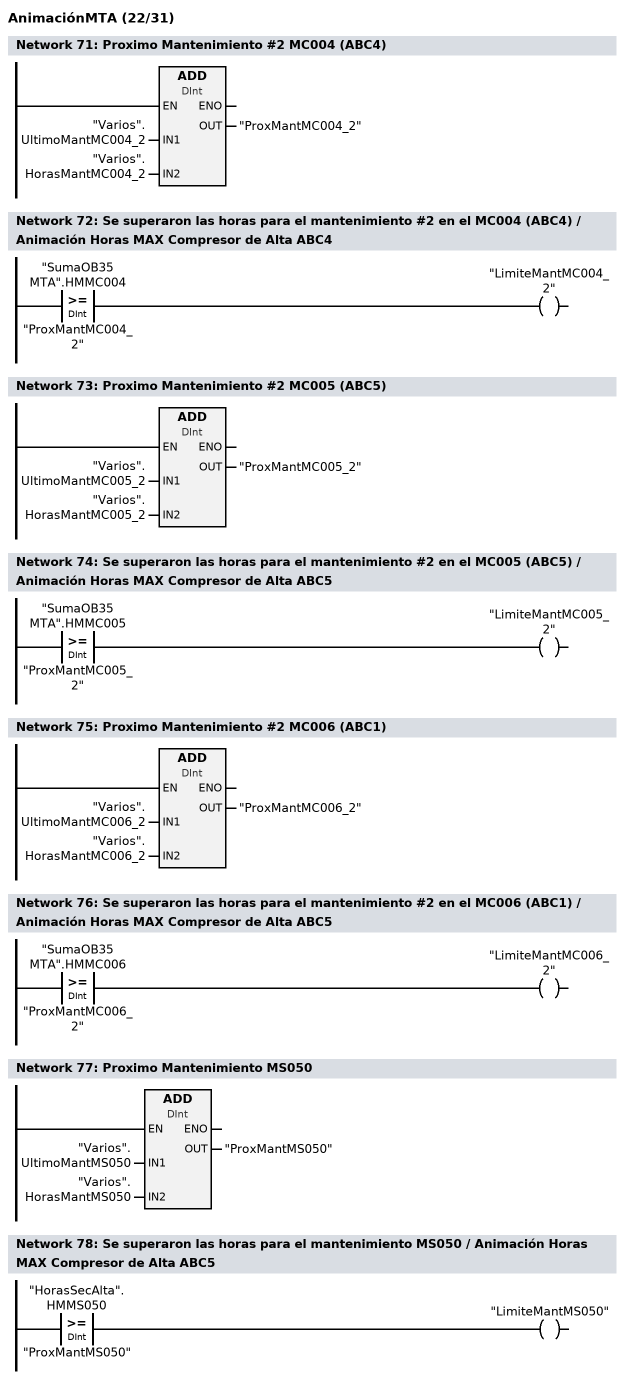
   RUNG wire#powerrail
      { S7_Templates := "SrcType := DInt"; S7_GenerateENO := "TRUE" } Add(in1 := "Varios".UltimoMantMC004_2, in2 := "Varios".HorasMantMC004_2, out => "ProxMantMC004_2")
   END_RUNG
   // the same network as SCL:
   "ProxMantMC004_2" := "Varios".UltimoMantMC004_2 + "Varios".HorasMantMC004_2;
END_REGION

REGION Network 72: Se superaron las horas para el mantenimiento #2 en el MC004 (ABC4) / Animación Horas MAX Compresor de Alta ABC4
   RUNG wire#powerrail
      { S7_Templates := "SrcType := DInt" } GE_Contact(in1 := "SumaOB35 MTA".HMMC004, in2 := "ProxMantMC004_2")
      Coil( "LimiteMantMC004_2" )
   END_RUNG
   // the same network as SCL:
   "LimiteMantMC004_2" := "SumaOB35 MTA".HMMC004 >= "ProxMantMC004_2";
END_REGION

REGION Network 73: Proximo Mantenimiento #2 MC005 (ABC5)
   RUNG wire#powerrail
      { S7_Templates := "SrcType := DInt"; S7_GenerateENO := "TRUE" } Add(in1 := "Varios".UltimoMantMC005_2, in2 := "Varios".HorasMantMC005_2, out => "ProxMantMC005_2")
   END_RUNG
   // the same network as SCL:
   "ProxMantMC005_2" := "Varios".UltimoMantMC005_2 + "Varios".HorasMantMC005_2;
END_REGION

REGION Network 74: Se superaron las horas para el mantenimiento #2 en el MC005 (ABC5) / Animación Horas MAX Compresor de Alta ABC5
   RUNG wire#powerrail
      { S7_Templates := "SrcType := DInt" } GE_Contact(in1 := "SumaOB35 MTA".HMMC005, in2 := "ProxMantMC005_2")
      Coil( "LimiteMantMC005_2" )
   END_RUNG
   // the same network as SCL:
   "LimiteMantMC005_2" := "SumaOB35 MTA".HMMC005 >= "ProxMantMC005_2";
END_REGION

REGION Network 75: Proximo Mantenimiento #2 MC006 (ABC1)
   RUNG wire#powerrail
      { S7_Templates := "SrcType := DInt"; S7_GenerateENO := "TRUE" } Add(in1 := "Varios".UltimoMantMC006_2, in2 := "Varios".HorasMantMC006_2, out => "ProxMantMC006_2")
   END_RUNG
   // the same network as SCL:
   "ProxMantMC006_2" := "Varios".UltimoMantMC006_2 + "Varios".HorasMantMC006_2;
END_REGION

REGION Network 76: Se superaron las horas para el mantenimiento #2 en el MC006 (ABC1) / Animación Horas MAX Compresor de Alta ABC5
   RUNG wire#powerrail
      { S7_Templates := "SrcType := DInt" } GE_Contact(in1 := "SumaOB35 MTA".HMMC006, in2 := "ProxMantMC006_2")
      Coil( "LimiteMantMC006_2" )
   END_RUNG
   // the same network as SCL:
   "LimiteMantMC006_2" := "SumaOB35 MTA".HMMC006 >= "ProxMantMC006_2";
END_REGION

REGION Network 77: Proximo Mantenimiento MS050
   RUNG wire#powerrail
      { S7_Templates := "SrcType := DInt"; S7_GenerateENO := "TRUE" } Add(in1 := "Varios".UltimoMantMS050, in2 := "Varios".HorasMantMS050, out => "ProxMantMS050")
   END_RUNG
   // the same network as SCL:
   "ProxMantMS050" := "Varios".UltimoMantMS050 + "Varios".HorasMantMS050;
END_REGION

REGION Network 78: Se superaron las horas para el mantenimiento MS050 / Animación Horas MAX Compresor de Alta ABC5
   RUNG wire#powerrail
      { S7_Templates := "SrcType := DInt" } GE_Contact(in1 := "HorasSecAlta".HMMS050, in2 := "ProxMantMS050")
      Coil( "LimiteMantMS050" )
   END_RUNG
   // the same network as SCL:
   "LimiteMantMS050" := "HorasSecAlta".HMMS050 >= "ProxMantMS050";
END_REGION

REGION Network 79: Proximo Mantenimiento MS051
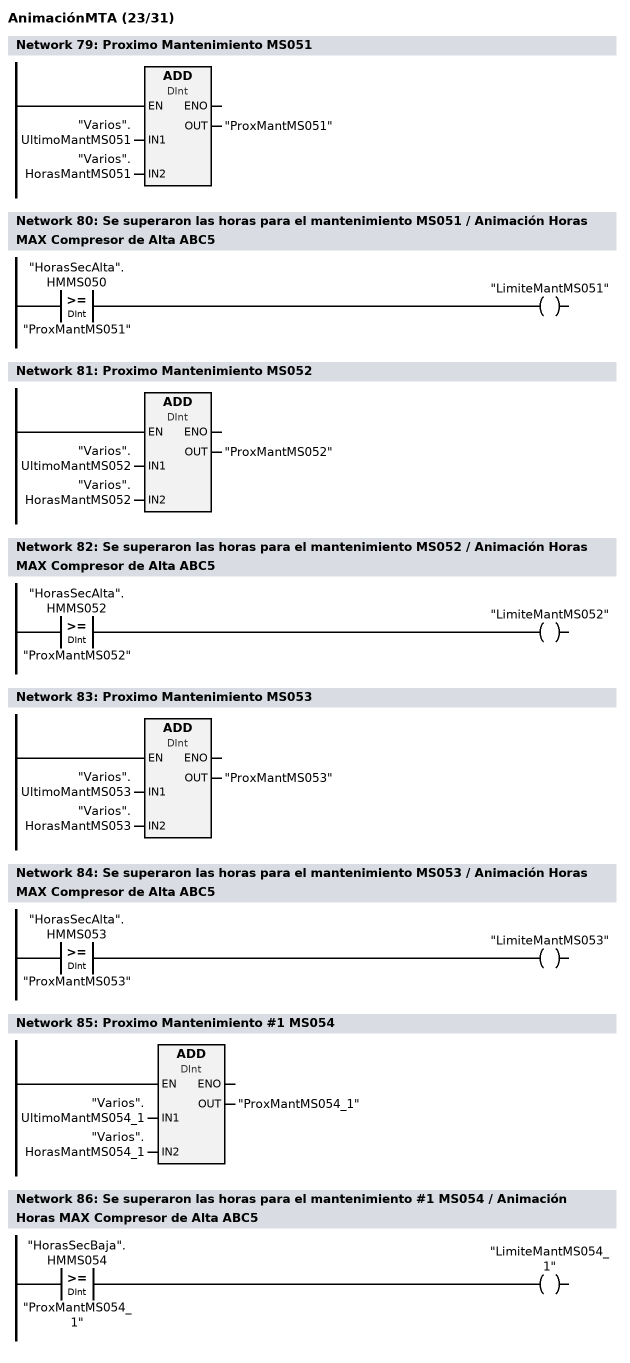
   RUNG wire#powerrail
      { S7_Templates := "SrcType := DInt"; S7_GenerateENO := "TRUE" } Add(in1 := "Varios".UltimoMantMS051, in2 := "Varios".HorasMantMS051, out => "ProxMantMS051")
   END_RUNG
   // the same network as SCL:
   "ProxMantMS051" := "Varios".UltimoMantMS051 + "Varios".HorasMantMS051;
END_REGION

REGION Network 80: Se superaron las horas para el mantenimiento MS051 / Animación Horas MAX Compresor de Alta ABC5
   RUNG wire#powerrail
      { S7_Templates := "SrcType := DInt" } GE_Contact(in1 := "HorasSecAlta".HMMS050, in2 := "ProxMantMS051")
      Coil( "LimiteMantMS051" )
   END_RUNG
   // the same network as SCL:
   "LimiteMantMS051" := "HorasSecAlta".HMMS050 >= "ProxMantMS051";
END_REGION

REGION Network 81: Proximo Mantenimiento MS052
   RUNG wire#powerrail
      { S7_Templates := "SrcType := DInt"; S7_GenerateENO := "TRUE" } Add(in1 := "Varios".UltimoMantMS052, in2 := "Varios".HorasMantMS052, out => "ProxMantMS052")
   END_RUNG
   // the same network as SCL:
   "ProxMantMS052" := "Varios".UltimoMantMS052 + "Varios".HorasMantMS052;
END_REGION

REGION Network 82: Se superaron las horas para el mantenimiento MS052 / Animación Horas MAX Compresor de Alta ABC5
   RUNG wire#powerrail
      { S7_Templates := "SrcType := DInt" } GE_Contact(in1 := "HorasSecAlta".HMMS052, in2 := "ProxMantMS052")
      Coil( "LimiteMantMS052" )
   END_RUNG
   // the same network as SCL:
   "LimiteMantMS052" := "HorasSecAlta".HMMS052 >= "ProxMantMS052";
END_REGION

REGION Network 83: Proximo Mantenimiento MS053
   RUNG wire#powerrail
      { S7_Templates := "SrcType := DInt"; S7_GenerateENO := "TRUE" } Add(in1 := "Varios".UltimoMantMS053, in2 := "Varios".HorasMantMS053, out => "ProxMantMS053")
   END_RUNG
   // the same network as SCL:
   "ProxMantMS053" := "Varios".UltimoMantMS053 + "Varios".HorasMantMS053;
END_REGION

REGION Network 84: Se superaron las horas para el mantenimiento MS053 / Animación Horas MAX Compresor de Alta ABC5
   RUNG wire#powerrail
      { S7_Templates := "SrcType := DInt" } GE_Contact(in1 := "HorasSecAlta".HMMS053, in2 := "ProxMantMS053")
      Coil( "LimiteMantMS053" )
   END_RUNG
   // the same network as SCL:
   "LimiteMantMS053" := "HorasSecAlta".HMMS053 >= "ProxMantMS053";
END_REGION

REGION Network 85: Proximo Mantenimiento #1 MS054
   RUNG wire#powerrail
      { S7_Templates := "SrcType := DInt"; S7_GenerateENO := "TRUE" } Add(in1 := "Varios".UltimoMantMS054_1, in2 := "Varios".HorasMantMS054_1, out => "ProxMantMS054_1")
   END_RUNG
   // the same network as SCL:
   "ProxMantMS054_1" := "Varios".UltimoMantMS054_1 + "Varios".HorasMantMS054_1;
END_REGION

REGION Network 86: Se superaron las horas para el mantenimiento #1 MS054 / Animación Horas MAX Compresor de Alta ABC5
   RUNG wire#powerrail
      { S7_Templates := "SrcType := DInt" } GE_Contact(in1 := "HorasSecBaja".HMMS054, in2 := "ProxMantMS054_1")
      Coil( "LimiteMantMS054_1" )
   END_RUNG
   // the same network as SCL:
   "LimiteMantMS054_1" := "HorasSecBaja".HMMS054 >= "ProxMantMS054_1";
END_REGION

REGION Network 87: Proximo Mantenimiento #2 MS054
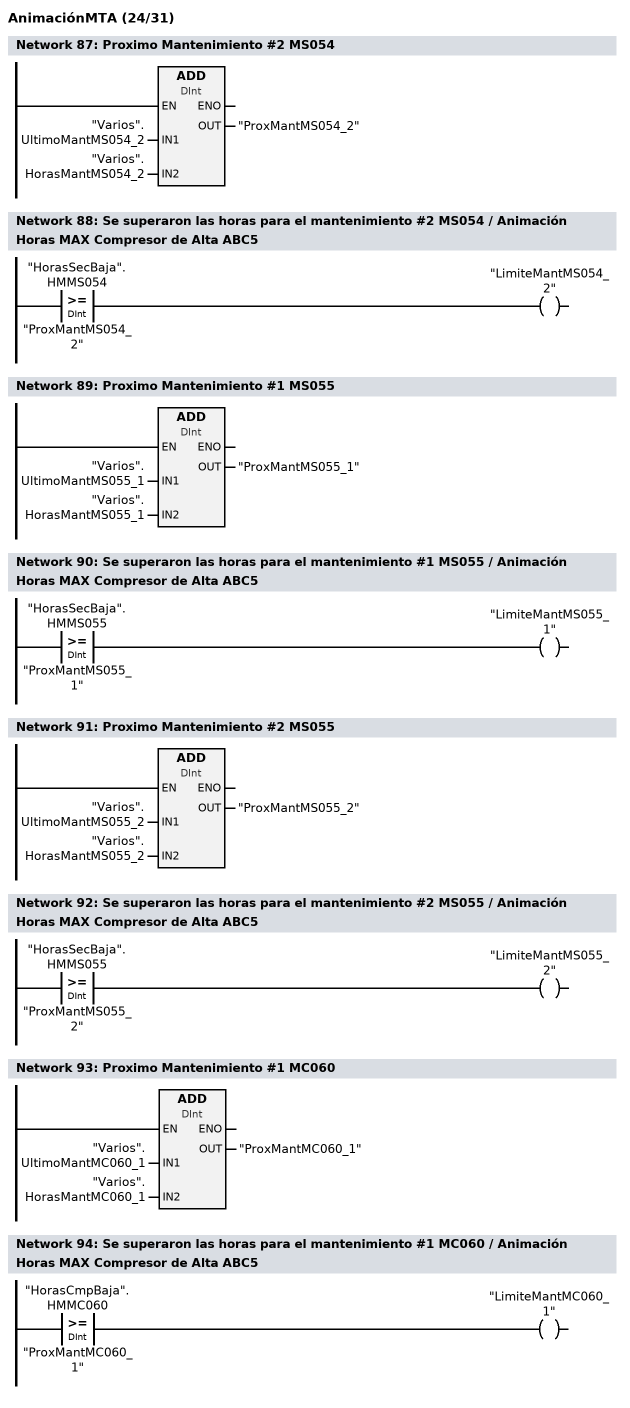
   RUNG wire#powerrail
      { S7_Templates := "SrcType := DInt"; S7_GenerateENO := "TRUE" } Add(in1 := "Varios".UltimoMantMS054_2, in2 := "Varios".HorasMantMS054_2, out => "ProxMantMS054_2")
   END_RUNG
   // the same network as SCL:
   "ProxMantMS054_2" := "Varios".UltimoMantMS054_2 + "Varios".HorasMantMS054_2;
END_REGION

REGION Network 88: Se superaron las horas para el mantenimiento #2 MS054 / Animación Horas MAX Compresor de Alta ABC5
   RUNG wire#powerrail
      { S7_Templates := "SrcType := DInt" } GE_Contact(in1 := "HorasSecBaja".HMMS054, in2 := "ProxMantMS054_2")
      Coil( "LimiteMantMS054_2" )
   END_RUNG
   // the same network as SCL:
   "LimiteMantMS054_2" := "HorasSecBaja".HMMS054 >= "ProxMantMS054_2";
END_REGION

REGION Network 89: Proximo Mantenimiento #1 MS055
   RUNG wire#powerrail
      { S7_Templates := "SrcType := DInt"; S7_GenerateENO := "TRUE" } Add(in1 := "Varios".UltimoMantMS055_1, in2 := "Varios".HorasMantMS055_1, out => "ProxMantMS055_1")
   END_RUNG
   // the same network as SCL:
   "ProxMantMS055_1" := "Varios".UltimoMantMS055_1 + "Varios".HorasMantMS055_1;
END_REGION

REGION Network 90: Se superaron las horas para el mantenimiento #1 MS055 / Animación Horas MAX Compresor de Alta ABC5
   RUNG wire#powerrail
      { S7_Templates := "SrcType := DInt" } GE_Contact(in1 := "HorasSecBaja".HMMS055, in2 := "ProxMantMS055_1")
      Coil( "LimiteMantMS055_1" )
   END_RUNG
   // the same network as SCL:
   "LimiteMantMS055_1" := "HorasSecBaja".HMMS055 >= "ProxMantMS055_1";
END_REGION

REGION Network 91: Proximo Mantenimiento #2 MS055
   RUNG wire#powerrail
      { S7_Templates := "SrcType := DInt"; S7_GenerateENO := "TRUE" } Add(in1 := "Varios".UltimoMantMS055_2, in2 := "Varios".HorasMantMS055_2, out => "ProxMantMS055_2")
   END_RUNG
   // the same network as SCL:
   "ProxMantMS055_2" := "Varios".UltimoMantMS055_2 + "Varios".HorasMantMS055_2;
END_REGION

REGION Network 92: Se superaron las horas para el mantenimiento #2 MS055 / Animación Horas MAX Compresor de Alta ABC5
   RUNG wire#powerrail
      { S7_Templates := "SrcType := DInt" } GE_Contact(in1 := "HorasSecBaja".HMMS055, in2 := "ProxMantMS055_2")
      Coil( "LimiteMantMS055_2" )
   END_RUNG
   // the same network as SCL:
   "LimiteMantMS055_2" := "HorasSecBaja".HMMS055 >= "ProxMantMS055_2";
END_REGION

REGION Network 93: Proximo Mantenimiento #1 MC060
   RUNG wire#powerrail
      { S7_Templates := "SrcType := DInt"; S7_GenerateENO := "TRUE" } Add(in1 := "Varios".UltimoMantMC060_1, in2 := "Varios".HorasMantMC060_1, out => "ProxMantMC060_1")
   END_RUNG
   // the same network as SCL:
   "ProxMantMC060_1" := "Varios".UltimoMantMC060_1 + "Varios".HorasMantMC060_1;
END_REGION

REGION Network 94: Se superaron las horas para el mantenimiento #1 MC060 / Animación Horas MAX Compresor de Alta ABC5
   RUNG wire#powerrail
      { S7_Templates := "SrcType := DInt" } GE_Contact(in1 := "HorasCmpBaja".HMMC060, in2 := "ProxMantMC060_1")
      Coil( "LimiteMantMC060_1" )
   END_RUNG
   // the same network as SCL:
   "LimiteMantMC060_1" := "HorasCmpBaja".HMMC060 >= "ProxMantMC060_1";
END_REGION

REGION Network 95: Proximo Mantenimiento #2 MC060
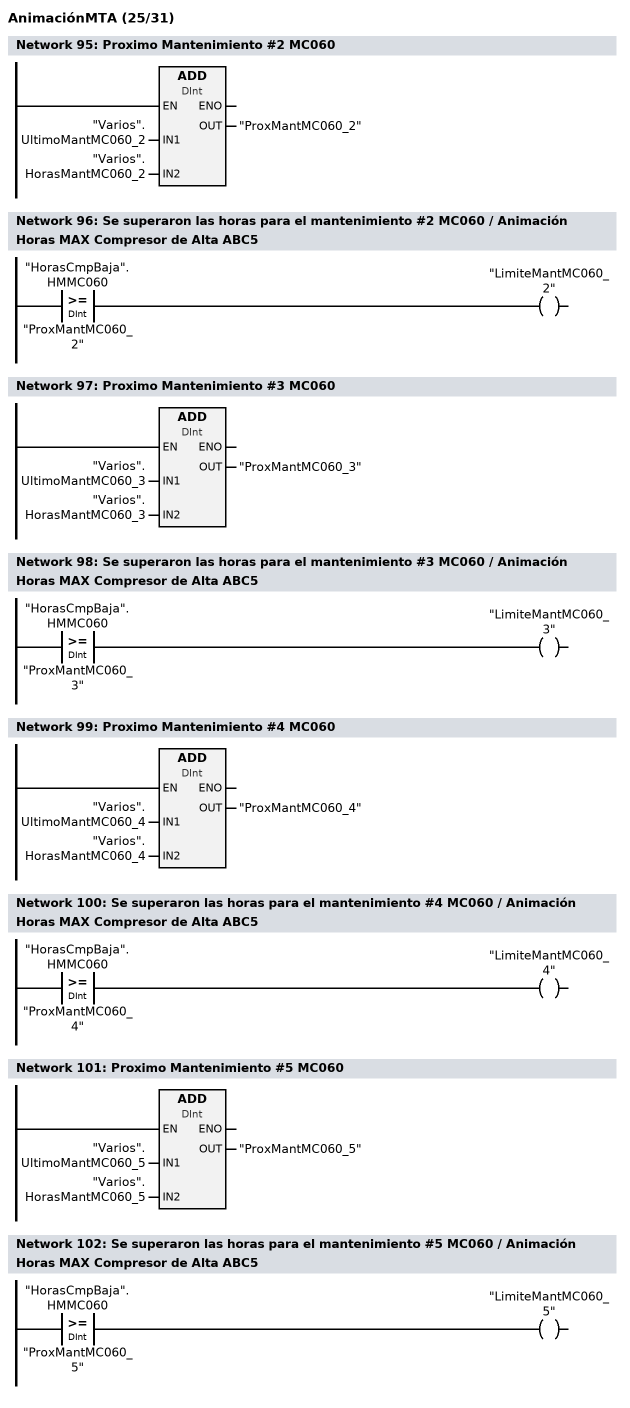
   RUNG wire#powerrail
      { S7_Templates := "SrcType := DInt"; S7_GenerateENO := "TRUE" } Add(in1 := "Varios".UltimoMantMC060_2, in2 := "Varios".HorasMantMC060_2, out => "ProxMantMC060_2")
   END_RUNG
   // the same network as SCL:
   "ProxMantMC060_2" := "Varios".UltimoMantMC060_2 + "Varios".HorasMantMC060_2;
END_REGION

REGION Network 96: Se superaron las horas para el mantenimiento #2 MC060 / Animación Horas MAX Compresor de Alta ABC5
   RUNG wire#powerrail
      { S7_Templates := "SrcType := DInt" } GE_Contact(in1 := "HorasCmpBaja".HMMC060, in2 := "ProxMantMC060_2")
      Coil( "LimiteMantMC060_2" )
   END_RUNG
   // the same network as SCL:
   "LimiteMantMC060_2" := "HorasCmpBaja".HMMC060 >= "ProxMantMC060_2";
END_REGION

REGION Network 97: Proximo Mantenimiento #3 MC060
   RUNG wire#powerrail
      { S7_Templates := "SrcType := DInt"; S7_GenerateENO := "TRUE" } Add(in1 := "Varios".UltimoMantMC060_3, in2 := "Varios".HorasMantMC060_3, out => "ProxMantMC060_3")
   END_RUNG
   // the same network as SCL:
   "ProxMantMC060_3" := "Varios".UltimoMantMC060_3 + "Varios".HorasMantMC060_3;
END_REGION

REGION Network 98: Se superaron las horas para el mantenimiento #3 MC060 / Animación Horas MAX Compresor de Alta ABC5
   RUNG wire#powerrail
      { S7_Templates := "SrcType := DInt" } GE_Contact(in1 := "HorasCmpBaja".HMMC060, in2 := "ProxMantMC060_3")
      Coil( "LimiteMantMC060_3" )
   END_RUNG
   // the same network as SCL:
   "LimiteMantMC060_3" := "HorasCmpBaja".HMMC060 >= "ProxMantMC060_3";
END_REGION

REGION Network 99: Proximo Mantenimiento #4 MC060
   RUNG wire#powerrail
      { S7_Templates := "SrcType := DInt"; S7_GenerateENO := "TRUE" } Add(in1 := "Varios".UltimoMantMC060_4, in2 := "Varios".HorasMantMC060_4, out => "ProxMantMC060_4")
   END_RUNG
   // the same network as SCL:
   "ProxMantMC060_4" := "Varios".UltimoMantMC060_4 + "Varios".HorasMantMC060_4;
END_REGION

REGION Network 100: Se superaron las horas para el mantenimiento #4 MC060 / Animación Horas MAX Compresor de Alta ABC5
   RUNG wire#powerrail
      { S7_Templates := "SrcType := DInt" } GE_Contact(in1 := "HorasCmpBaja".HMMC060, in2 := "ProxMantMC060_4")
      Coil( "LimiteMantMC060_4" )
   END_RUNG
   // the same network as SCL:
   "LimiteMantMC060_4" := "HorasCmpBaja".HMMC060 >= "ProxMantMC060_4";
END_REGION

REGION Network 101: Proximo Mantenimiento #5 MC060
   RUNG wire#powerrail
      { S7_Templates := "SrcType := DInt"; S7_GenerateENO := "TRUE" } Add(in1 := "Varios".UltimoMantMC060_5, in2 := "Varios".HorasMantMC060_5, out => "ProxMantMC060_5")
   END_RUNG
   // the same network as SCL:
   "ProxMantMC060_5" := "Varios".UltimoMantMC060_5 + "Varios".HorasMantMC060_5;
END_REGION

REGION Network 102: Se superaron las horas para el mantenimiento #5 MC060 / Animación Horas MAX Compresor de Alta ABC5
   RUNG wire#powerrail
      { S7_Templates := "SrcType := DInt" } GE_Contact(in1 := "HorasCmpBaja".HMMC060, in2 := "ProxMantMC060_5")
      Coil( "LimiteMantMC060_5" )
   END_RUNG
   // the same network as SCL:
   "LimiteMantMC060_5" := "HorasCmpBaja".HMMC060 >= "ProxMantMC060_5";
END_REGION

REGION Network 103: Proximo Mantenimiento #1 MC061
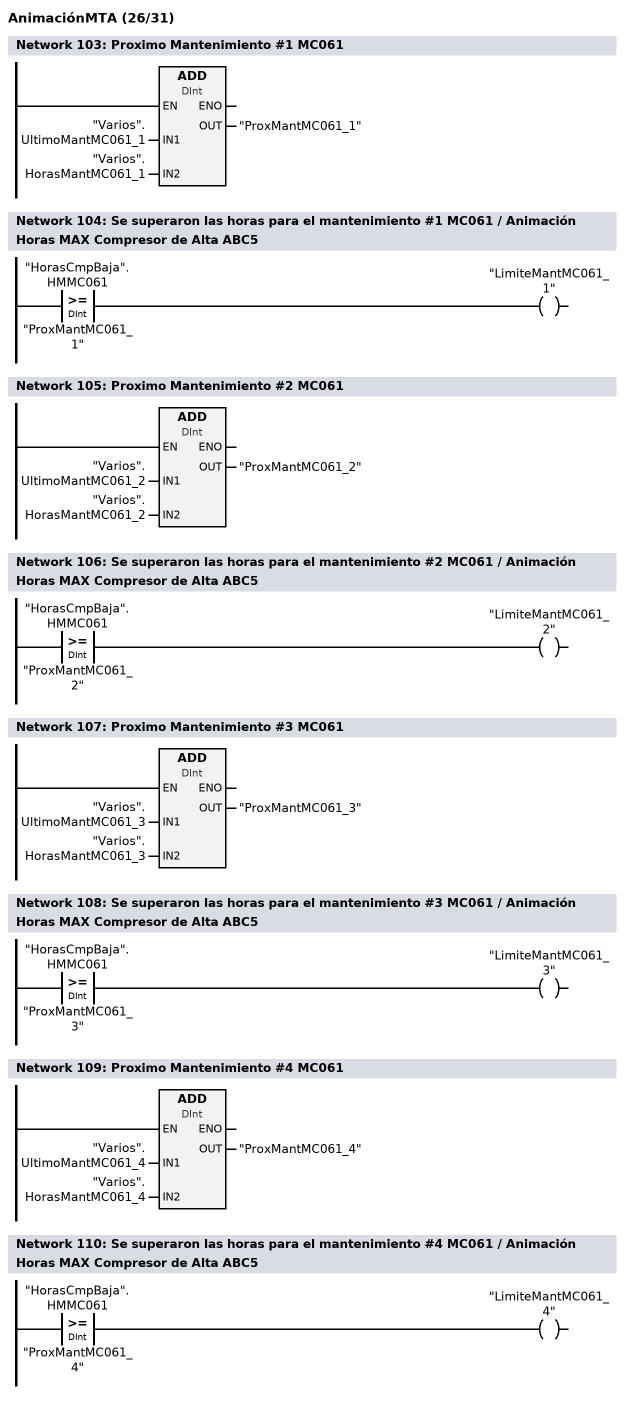
   RUNG wire#powerrail
      { S7_Templates := "SrcType := DInt"; S7_GenerateENO := "TRUE" } Add(in1 := "Varios".UltimoMantMC061_1, in2 := "Varios".HorasMantMC061_1, out => "ProxMantMC061_1")
   END_RUNG
   // the same network as SCL:
   "ProxMantMC061_1" := "Varios".UltimoMantMC061_1 + "Varios".HorasMantMC061_1;
END_REGION

REGION Network 104: Se superaron las horas para el mantenimiento #1 MC061 / Animación Horas MAX Compresor de Alta ABC5
   RUNG wire#powerrail
      { S7_Templates := "SrcType := DInt" } GE_Contact(in1 := "HorasCmpBaja".HMMC061, in2 := "ProxMantMC061_1")
      Coil( "LimiteMantMC061_1" )
   END_RUNG
   // the same network as SCL:
   "LimiteMantMC061_1" := "HorasCmpBaja".HMMC061 >= "ProxMantMC061_1";
END_REGION

REGION Network 105: Proximo Mantenimiento #2 MC061
   RUNG wire#powerrail
      { S7_Templates := "SrcType := DInt"; S7_GenerateENO := "TRUE" } Add(in1 := "Varios".UltimoMantMC061_2, in2 := "Varios".HorasMantMC061_2, out => "ProxMantMC061_2")
   END_RUNG
   // the same network as SCL:
   "ProxMantMC061_2" := "Varios".UltimoMantMC061_2 + "Varios".HorasMantMC061_2;
END_REGION

REGION Network 106: Se superaron las horas para el mantenimiento #2 MC061 / Animación Horas MAX Compresor de Alta ABC5
   RUNG wire#powerrail
      { S7_Templates := "SrcType := DInt" } GE_Contact(in1 := "HorasCmpBaja".HMMC061, in2 := "ProxMantMC061_2")
      Coil( "LimiteMantMC061_2" )
   END_RUNG
   // the same network as SCL:
   "LimiteMantMC061_2" := "HorasCmpBaja".HMMC061 >= "ProxMantMC061_2";
END_REGION

REGION Network 107: Proximo Mantenimiento #3 MC061
   RUNG wire#powerrail
      { S7_Templates := "SrcType := DInt"; S7_GenerateENO := "TRUE" } Add(in1 := "Varios".UltimoMantMC061_3, in2 := "Varios".HorasMantMC061_3, out => "ProxMantMC061_3")
   END_RUNG
   // the same network as SCL:
   "ProxMantMC061_3" := "Varios".UltimoMantMC061_3 + "Varios".HorasMantMC061_3;
END_REGION

REGION Network 108: Se superaron las horas para el mantenimiento #3 MC061 / Animación Horas MAX Compresor de Alta ABC5
   RUNG wire#powerrail
      { S7_Templates := "SrcType := DInt" } GE_Contact(in1 := "HorasCmpBaja".HMMC061, in2 := "ProxMantMC061_3")
      Coil( "LimiteMantMC061_3" )
   END_RUNG
   // the same network as SCL:
   "LimiteMantMC061_3" := "HorasCmpBaja".HMMC061 >= "ProxMantMC061_3";
END_REGION

REGION Network 109: Proximo Mantenimiento #4 MC061
   RUNG wire#powerrail
      { S7_Templates := "SrcType := DInt"; S7_GenerateENO := "TRUE" } Add(in1 := "Varios".UltimoMantMC061_4, in2 := "Varios".HorasMantMC061_4, out => "ProxMantMC061_4")
   END_RUNG
   // the same network as SCL:
   "ProxMantMC061_4" := "Varios".UltimoMantMC061_4 + "Varios".HorasMantMC061_4;
END_REGION

REGION Network 110: Se superaron las horas para el mantenimiento #4 MC061 / Animación Horas MAX Compresor de Alta ABC5
   RUNG wire#powerrail
      { S7_Templates := "SrcType := DInt" } GE_Contact(in1 := "HorasCmpBaja".HMMC061, in2 := "ProxMantMC061_4")
      Coil( "LimiteMantMC061_4" )
   END_RUNG
   // the same network as SCL:
   "LimiteMantMC061_4" := "HorasCmpBaja".HMMC061 >= "ProxMantMC061_4";
END_REGION

REGION Network 111: Proximo Mantenimiento #5 MC061
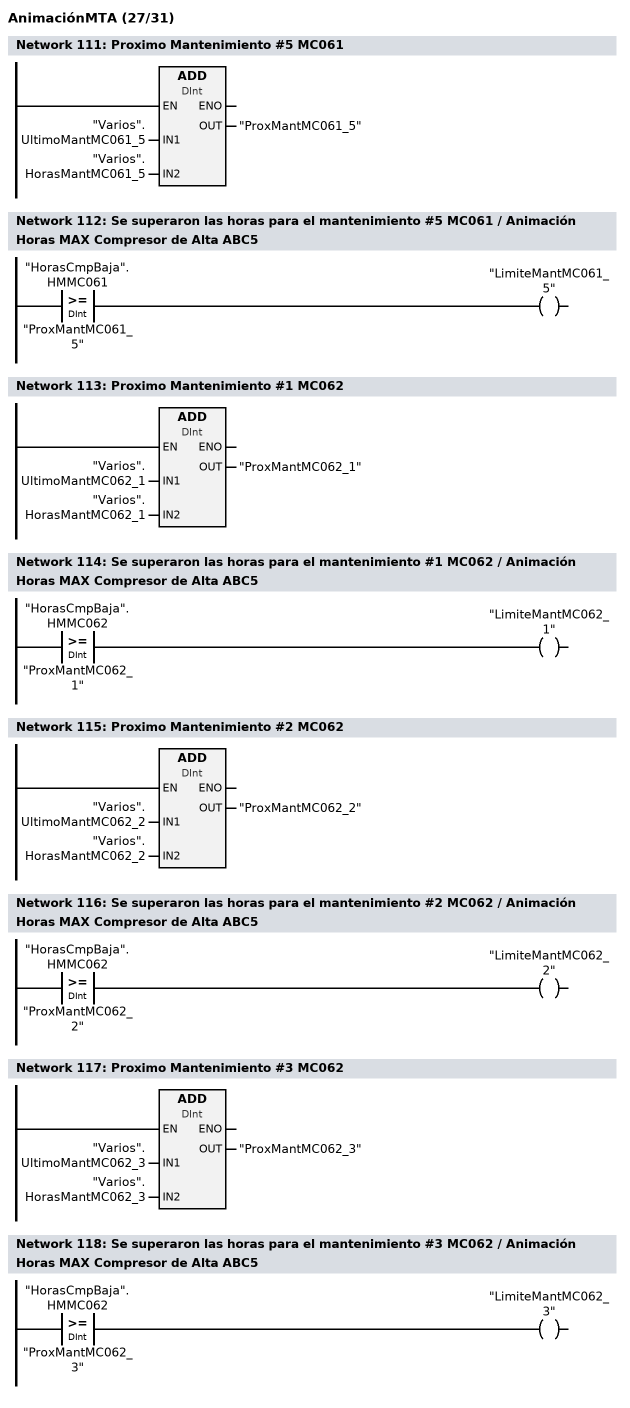
   RUNG wire#powerrail
      { S7_Templates := "SrcType := DInt"; S7_GenerateENO := "TRUE" } Add(in1 := "Varios".UltimoMantMC061_5, in2 := "Varios".HorasMantMC061_5, out => "ProxMantMC061_5")
   END_RUNG
   // the same network as SCL:
   "ProxMantMC061_5" := "Varios".UltimoMantMC061_5 + "Varios".HorasMantMC061_5;
END_REGION

REGION Network 112: Se superaron las horas para el mantenimiento #5 MC061 / Animación Horas MAX Compresor de Alta ABC5
   RUNG wire#powerrail
      { S7_Templates := "SrcType := DInt" } GE_Contact(in1 := "HorasCmpBaja".HMMC061, in2 := "ProxMantMC061_5")
      Coil( "LimiteMantMC061_5" )
   END_RUNG
   // the same network as SCL:
   "LimiteMantMC061_5" := "HorasCmpBaja".HMMC061 >= "ProxMantMC061_5";
END_REGION

REGION Network 113: Proximo Mantenimiento #1 MC062
   RUNG wire#powerrail
      { S7_Templates := "SrcType := DInt"; S7_GenerateENO := "TRUE" } Add(in1 := "Varios".UltimoMantMC062_1, in2 := "Varios".HorasMantMC062_1, out => "ProxMantMC062_1")
   END_RUNG
   // the same network as SCL:
   "ProxMantMC062_1" := "Varios".UltimoMantMC062_1 + "Varios".HorasMantMC062_1;
END_REGION

REGION Network 114: Se superaron las horas para el mantenimiento #1 MC062 / Animación Horas MAX Compresor de Alta ABC5
   RUNG wire#powerrail
      { S7_Templates := "SrcType := DInt" } GE_Contact(in1 := "HorasCmpBaja".HMMC062, in2 := "ProxMantMC062_1")
      Coil( "LimiteMantMC062_1" )
   END_RUNG
   // the same network as SCL:
   "LimiteMantMC062_1" := "HorasCmpBaja".HMMC062 >= "ProxMantMC062_1";
END_REGION

REGION Network 115: Proximo Mantenimiento #2 MC062
   RUNG wire#powerrail
      { S7_Templates := "SrcType := DInt"; S7_GenerateENO := "TRUE" } Add(in1 := "Varios".UltimoMantMC062_2, in2 := "Varios".HorasMantMC062_2, out => "ProxMantMC062_2")
   END_RUNG
   // the same network as SCL:
   "ProxMantMC062_2" := "Varios".UltimoMantMC062_2 + "Varios".HorasMantMC062_2;
END_REGION

REGION Network 116: Se superaron las horas para el mantenimiento #2 MC062 / Animación Horas MAX Compresor de Alta ABC5
   RUNG wire#powerrail
      { S7_Templates := "SrcType := DInt" } GE_Contact(in1 := "HorasCmpBaja".HMMC062, in2 := "ProxMantMC062_2")
      Coil( "LimiteMantMC062_2" )
   END_RUNG
   // the same network as SCL:
   "LimiteMantMC062_2" := "HorasCmpBaja".HMMC062 >= "ProxMantMC062_2";
END_REGION

REGION Network 117: Proximo Mantenimiento #3 MC062
   RUNG wire#powerrail
      { S7_Templates := "SrcType := DInt"; S7_GenerateENO := "TRUE" } Add(in1 := "Varios".UltimoMantMC062_3, in2 := "Varios".HorasMantMC062_3, out => "ProxMantMC062_3")
   END_RUNG
   // the same network as SCL:
   "ProxMantMC062_3" := "Varios".UltimoMantMC062_3 + "Varios".HorasMantMC062_3;
END_REGION

REGION Network 118: Se superaron las horas para el mantenimiento #3 MC062 / Animación Horas MAX Compresor de Alta ABC5
   RUNG wire#powerrail
      { S7_Templates := "SrcType := DInt" } GE_Contact(in1 := "HorasCmpBaja".HMMC062, in2 := "ProxMantMC062_3")
      Coil( "LimiteMantMC062_3" )
   END_RUNG
   // the same network as SCL:
   "LimiteMantMC062_3" := "HorasCmpBaja".HMMC062 >= "ProxMantMC062_3";
END_REGION

REGION Network 119: Proximo Mantenimiento #4 MC062
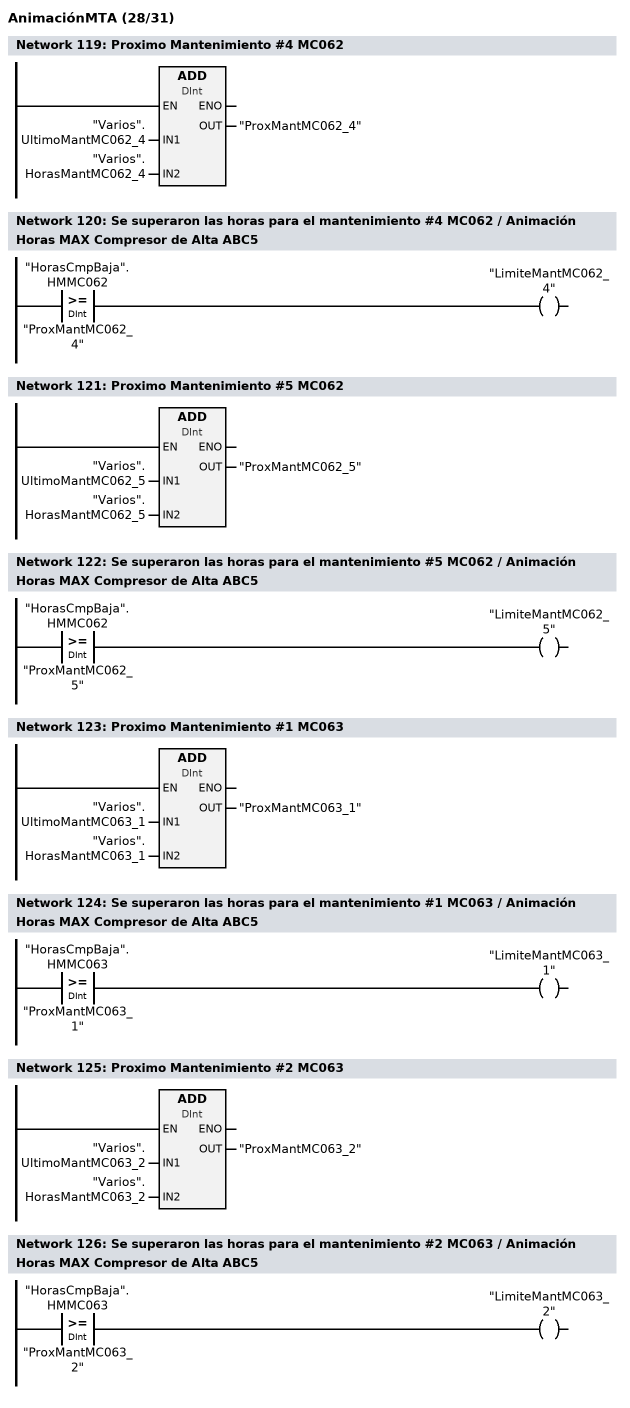
   RUNG wire#powerrail
      { S7_Templates := "SrcType := DInt"; S7_GenerateENO := "TRUE" } Add(in1 := "Varios".UltimoMantMC062_4, in2 := "Varios".HorasMantMC062_4, out => "ProxMantMC062_4")
   END_RUNG
   // the same network as SCL:
   "ProxMantMC062_4" := "Varios".UltimoMantMC062_4 + "Varios".HorasMantMC062_4;
END_REGION

REGION Network 120: Se superaron las horas para el mantenimiento #4 MC062 / Animación Horas MAX Compresor de Alta ABC5
   RUNG wire#powerrail
      { S7_Templates := "SrcType := DInt" } GE_Contact(in1 := "HorasCmpBaja".HMMC062, in2 := "ProxMantMC062_4")
      Coil( "LimiteMantMC062_4" )
   END_RUNG
   // the same network as SCL:
   "LimiteMantMC062_4" := "HorasCmpBaja".HMMC062 >= "ProxMantMC062_4";
END_REGION

REGION Network 121: Proximo Mantenimiento #5 MC062
   RUNG wire#powerrail
      { S7_Templates := "SrcType := DInt"; S7_GenerateENO := "TRUE" } Add(in1 := "Varios".UltimoMantMC062_5, in2 := "Varios".HorasMantMC062_5, out => "ProxMantMC062_5")
   END_RUNG
   // the same network as SCL:
   "ProxMantMC062_5" := "Varios".UltimoMantMC062_5 + "Varios".HorasMantMC062_5;
END_REGION

REGION Network 122: Se superaron las horas para el mantenimiento #5 MC062 / Animación Horas MAX Compresor de Alta ABC5
   RUNG wire#powerrail
      { S7_Templates := "SrcType := DInt" } GE_Contact(in1 := "HorasCmpBaja".HMMC062, in2 := "ProxMantMC062_5")
      Coil( "LimiteMantMC062_5" )
   END_RUNG
   // the same network as SCL:
   "LimiteMantMC062_5" := "HorasCmpBaja".HMMC062 >= "ProxMantMC062_5";
END_REGION

REGION Network 123: Proximo Mantenimiento #1 MC063
   RUNG wire#powerrail
      { S7_Templates := "SrcType := DInt"; S7_GenerateENO := "TRUE" } Add(in1 := "Varios".UltimoMantMC063_1, in2 := "Varios".HorasMantMC063_1, out => "ProxMantMC063_1")
   END_RUNG
   // the same network as SCL:
   "ProxMantMC063_1" := "Varios".UltimoMantMC063_1 + "Varios".HorasMantMC063_1;
END_REGION

REGION Network 124: Se superaron las horas para el mantenimiento #1 MC063 / Animación Horas MAX Compresor de Alta ABC5
   RUNG wire#powerrail
      { S7_Templates := "SrcType := DInt" } GE_Contact(in1 := "HorasCmpBaja".HMMC063, in2 := "ProxMantMC063_1")
      Coil( "LimiteMantMC063_1" )
   END_RUNG
   // the same network as SCL:
   "LimiteMantMC063_1" := "HorasCmpBaja".HMMC063 >= "ProxMantMC063_1";
END_REGION

REGION Network 125: Proximo Mantenimiento #2 MC063
   RUNG wire#powerrail
      { S7_Templates := "SrcType := DInt"; S7_GenerateENO := "TRUE" } Add(in1 := "Varios".UltimoMantMC063_2, in2 := "Varios".HorasMantMC063_2, out => "ProxMantMC063_2")
   END_RUNG
   // the same network as SCL:
   "ProxMantMC063_2" := "Varios".UltimoMantMC063_2 + "Varios".HorasMantMC063_2;
END_REGION

REGION Network 126: Se superaron las horas para el mantenimiento #2 MC063 / Animación Horas MAX Compresor de Alta ABC5
   RUNG wire#powerrail
      { S7_Templates := "SrcType := DInt" } GE_Contact(in1 := "HorasCmpBaja".HMMC063, in2 := "ProxMantMC063_2")
      Coil( "LimiteMantMC063_2" )
   END_RUNG
   // the same network as SCL:
   "LimiteMantMC063_2" := "HorasCmpBaja".HMMC063 >= "ProxMantMC063_2";
END_REGION

REGION Network 127: Proximo Mantenimiento #3 MC063
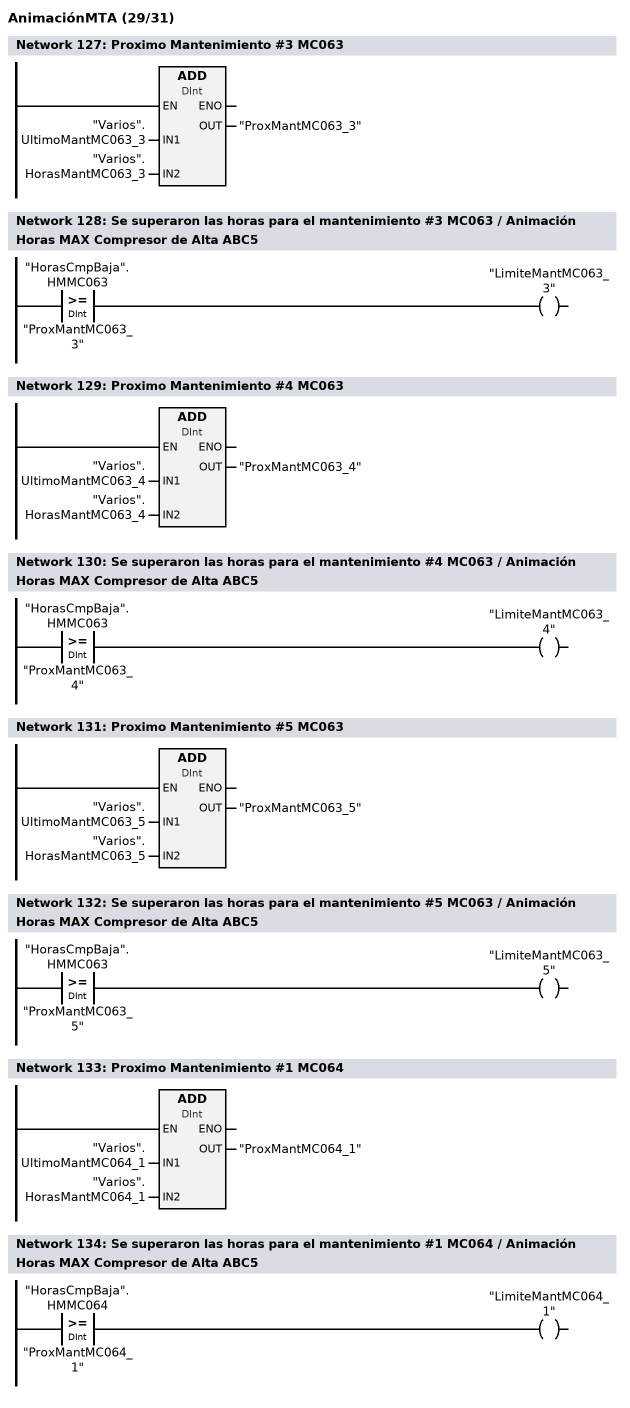
   RUNG wire#powerrail
      { S7_Templates := "SrcType := DInt"; S7_GenerateENO := "TRUE" } Add(in1 := "Varios".UltimoMantMC063_3, in2 := "Varios".HorasMantMC063_3, out => "ProxMantMC063_3")
   END_RUNG
   // the same network as SCL:
   "ProxMantMC063_3" := "Varios".UltimoMantMC063_3 + "Varios".HorasMantMC063_3;
END_REGION

REGION Network 128: Se superaron las horas para el mantenimiento #3 MC063 / Animación Horas MAX Compresor de Alta ABC5
   RUNG wire#powerrail
      { S7_Templates := "SrcType := DInt" } GE_Contact(in1 := "HorasCmpBaja".HMMC063, in2 := "ProxMantMC063_3")
      Coil( "LimiteMantMC063_3" )
   END_RUNG
   // the same network as SCL:
   "LimiteMantMC063_3" := "HorasCmpBaja".HMMC063 >= "ProxMantMC063_3";
END_REGION

REGION Network 129: Proximo Mantenimiento #4 MC063
   RUNG wire#powerrail
      { S7_Templates := "SrcType := DInt"; S7_GenerateENO := "TRUE" } Add(in1 := "Varios".UltimoMantMC063_4, in2 := "Varios".HorasMantMC063_4, out => "ProxMantMC063_4")
   END_RUNG
   // the same network as SCL:
   "ProxMantMC063_4" := "Varios".UltimoMantMC063_4 + "Varios".HorasMantMC063_4;
END_REGION

REGION Network 130: Se superaron las horas para el mantenimiento #4 MC063 / Animación Horas MAX Compresor de Alta ABC5
   RUNG wire#powerrail
      { S7_Templates := "SrcType := DInt" } GE_Contact(in1 := "HorasCmpBaja".HMMC063, in2 := "ProxMantMC063_4")
      Coil( "LimiteMantMC063_4" )
   END_RUNG
   // the same network as SCL:
   "LimiteMantMC063_4" := "HorasCmpBaja".HMMC063 >= "ProxMantMC063_4";
END_REGION

REGION Network 131: Proximo Mantenimiento #5 MC063
   RUNG wire#powerrail
      { S7_Templates := "SrcType := DInt"; S7_GenerateENO := "TRUE" } Add(in1 := "Varios".UltimoMantMC063_5, in2 := "Varios".HorasMantMC063_5, out => "ProxMantMC063_5")
   END_RUNG
   // the same network as SCL:
   "ProxMantMC063_5" := "Varios".UltimoMantMC063_5 + "Varios".HorasMantMC063_5;
END_REGION

REGION Network 132: Se superaron las horas para el mantenimiento #5 MC063 / Animación Horas MAX Compresor de Alta ABC5
   RUNG wire#powerrail
      { S7_Templates := "SrcType := DInt" } GE_Contact(in1 := "HorasCmpBaja".HMMC063, in2 := "ProxMantMC063_5")
      Coil( "LimiteMantMC063_5" )
   END_RUNG
   // the same network as SCL:
   "LimiteMantMC063_5" := "HorasCmpBaja".HMMC063 >= "ProxMantMC063_5";
END_REGION

REGION Network 133: Proximo Mantenimiento #1 MC064
   RUNG wire#powerrail
      { S7_Templates := "SrcType := DInt"; S7_GenerateENO := "TRUE" } Add(in1 := "Varios".UltimoMantMC064_1, in2 := "Varios".HorasMantMC064_1, out => "ProxMantMC064_1")
   END_RUNG
   // the same network as SCL:
   "ProxMantMC064_1" := "Varios".UltimoMantMC064_1 + "Varios".HorasMantMC064_1;
END_REGION

REGION Network 134: Se superaron las horas para el mantenimiento #1 MC064 / Animación Horas MAX Compresor de Alta ABC5
   RUNG wire#powerrail
      { S7_Templates := "SrcType := DInt" } GE_Contact(in1 := "HorasCmpBaja".HMMC064, in2 := "ProxMantMC064_1")
      Coil( "LimiteMantMC064_1" )
   END_RUNG
   // the same network as SCL:
   "LimiteMantMC064_1" := "HorasCmpBaja".HMMC064 >= "ProxMantMC064_1";
END_REGION

REGION Network 135: Proximo Mantenimiento #2 MC064
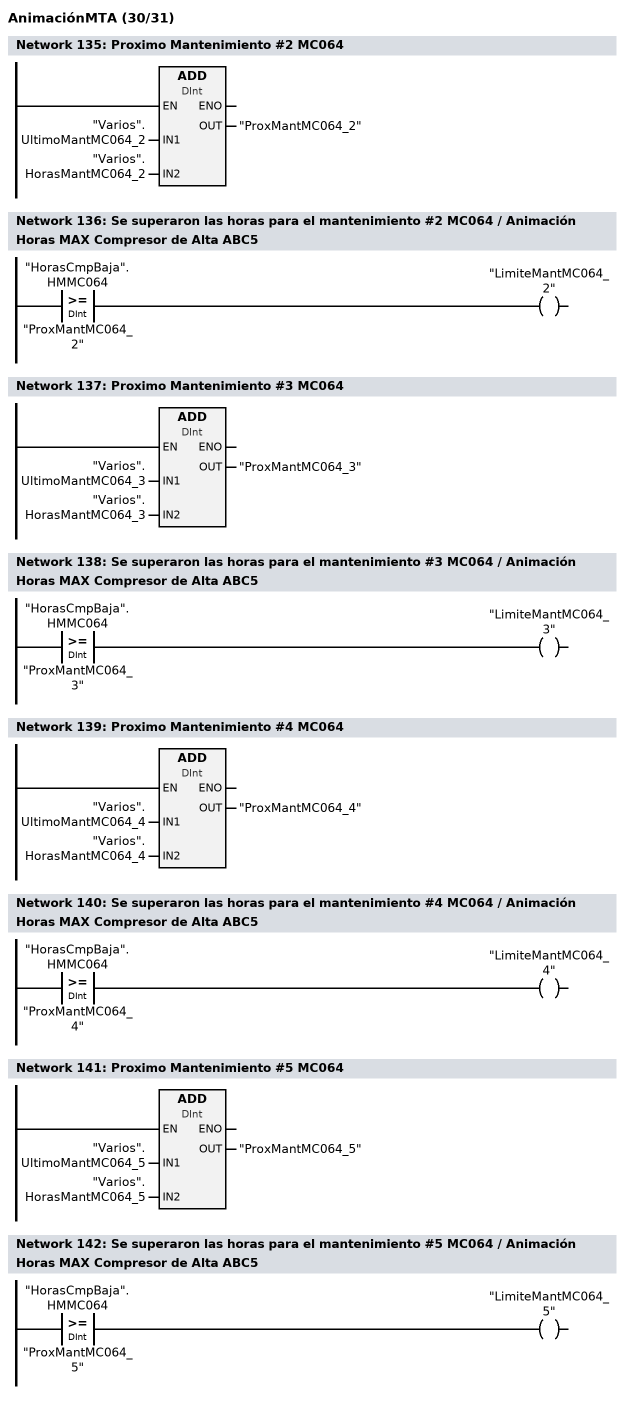
   RUNG wire#powerrail
      { S7_Templates := "SrcType := DInt"; S7_GenerateENO := "TRUE" } Add(in1 := "Varios".UltimoMantMC064_2, in2 := "Varios".HorasMantMC064_2, out => "ProxMantMC064_2")
   END_RUNG
   // the same network as SCL:
   "ProxMantMC064_2" := "Varios".UltimoMantMC064_2 + "Varios".HorasMantMC064_2;
END_REGION

REGION Network 136: Se superaron las horas para el mantenimiento #2 MC064 / Animación Horas MAX Compresor de Alta ABC5
   RUNG wire#powerrail
      { S7_Templates := "SrcType := DInt" } GE_Contact(in1 := "HorasCmpBaja".HMMC064, in2 := "ProxMantMC064_2")
      Coil( "LimiteMantMC064_2" )
   END_RUNG
   // the same network as SCL:
   "LimiteMantMC064_2" := "HorasCmpBaja".HMMC064 >= "ProxMantMC064_2";
END_REGION

REGION Network 137: Proximo Mantenimiento #3 MC064
   RUNG wire#powerrail
      { S7_Templates := "SrcType := DInt"; S7_GenerateENO := "TRUE" } Add(in1 := "Varios".UltimoMantMC064_3, in2 := "Varios".HorasMantMC064_3, out => "ProxMantMC064_3")
   END_RUNG
   // the same network as SCL:
   "ProxMantMC064_3" := "Varios".UltimoMantMC064_3 + "Varios".HorasMantMC064_3;
END_REGION

REGION Network 138: Se superaron las horas para el mantenimiento #3 MC064 / Animación Horas MAX Compresor de Alta ABC5
   RUNG wire#powerrail
      { S7_Templates := "SrcType := DInt" } GE_Contact(in1 := "HorasCmpBaja".HMMC064, in2 := "ProxMantMC064_3")
      Coil( "LimiteMantMC064_3" )
   END_RUNG
   // the same network as SCL:
   "LimiteMantMC064_3" := "HorasCmpBaja".HMMC064 >= "ProxMantMC064_3";
END_REGION

REGION Network 139: Proximo Mantenimiento #4 MC064
   RUNG wire#powerrail
      { S7_Templates := "SrcType := DInt"; S7_GenerateENO := "TRUE" } Add(in1 := "Varios".UltimoMantMC064_4, in2 := "Varios".HorasMantMC064_4, out => "ProxMantMC064_4")
   END_RUNG
   // the same network as SCL:
   "ProxMantMC064_4" := "Varios".UltimoMantMC064_4 + "Varios".HorasMantMC064_4;
END_REGION

REGION Network 140: Se superaron las horas para el mantenimiento #4 MC064 / Animación Horas MAX Compresor de Alta ABC5
   RUNG wire#powerrail
      { S7_Templates := "SrcType := DInt" } GE_Contact(in1 := "HorasCmpBaja".HMMC064, in2 := "ProxMantMC064_4")
      Coil( "LimiteMantMC064_4" )
   END_RUNG
   // the same network as SCL:
   "LimiteMantMC064_4" := "HorasCmpBaja".HMMC064 >= "ProxMantMC064_4";
END_REGION

REGION Network 141: Proximo Mantenimiento #5 MC064
   RUNG wire#powerrail
      { S7_Templates := "SrcType := DInt"; S7_GenerateENO := "TRUE" } Add(in1 := "Varios".UltimoMantMC064_5, in2 := "Varios".HorasMantMC064_5, out => "ProxMantMC064_5")
   END_RUNG
   // the same network as SCL:
   "ProxMantMC064_5" := "Varios".UltimoMantMC064_5 + "Varios".HorasMantMC064_5;
END_REGION

REGION Network 142: Se superaron las horas para el mantenimiento #5 MC064 / Animación Horas MAX Compresor de Alta ABC5
   RUNG wire#powerrail
      { S7_Templates := "SrcType := DInt" } GE_Contact(in1 := "HorasCmpBaja".HMMC064, in2 := "ProxMantMC064_5")
      Coil( "LimiteMantMC064_5" )
   END_RUNG
   // the same network as SCL:
   "LimiteMantMC064_5" := "HorasCmpBaja".HMMC064 >= "ProxMantMC064_5";
END_REGION

REGION Network 143: Próximo Mantenimento Booster 1
